(* Logix 5000 project; controller PLC_MCC1201_220AP1 vendor 1 type 14 code 164 rev 35.11; software revision 35.00; part 16 of 25 *)
(* tags used below, declared in another part *)
   AFI : ALIAS FOR B3[7].15;
   B151 : DINT[20];
   B152 : DINT[50];
   B153 : DINT[20];
   B154 : DINT[20];
   B155 : DINT[20];
   B3 : DINT[102];
   BT41_006 : MESSAGE;   // Block Transfer Read Control for Analog Input Card in Washer Panel
   BT41_007 : MESSAGE;   // Block Transfer Write Control for Analog Input Card in Washer Panel
   C1_ACK : ALIAS FOR N54[260].14;
   C1_ACTIVE_LAMP : ALIAS FOR N54[260].0;
   C1_BEACON : ALIAS FOR O[27].6;
   C1_BEACON2 : ALIAS FOR O[47].10;
   C1_HORN : ALIAS FOR O[27].5;
   C1_NTH_IN_LMP : ALIAS FOR N54[260].10;
   C1_NTH_IN_PE : ALIAS FOR N54[260].6;
   C1_NTH_IN_SS : ALIAS FOR N54[260].2;
   C1_NTH_OUT_LMP : ALIAS FOR N54[260].9;
   C1_NTH_OUT_PE : ALIAS FOR N54[260].5;
   C1_NTH_OUT_SS : ALIAS FOR N54[260].1;
   C1_STH_IN_LMP : ALIAS FOR N54[260].12;
   C1_STH_IN_PE : ALIAS FOR N54[260].8;
   C1_STH_IN_SS : ALIAS FOR N54[260].4;
   C1_STH_OUT_LMP : ALIAS FOR N54[260].11;
   C1_STH_OUT_PE : ALIAS FOR N54[260].7;
   C1_STH_OUT_SS : ALIAS FOR N54[260].3;
   C2_ACTIVE_LAMP : ALIAS FOR N54[261].0;
   C2_NTH_IN_LMP : ALIAS FOR N54[261].10;
   C2_NTH_IN_PE : ALIAS FOR N54[261].6;
   C2_NTH_IN_SS : ALIAS FOR N54[261].2;
   C2_NTH_OUT_LMP : ALIAS FOR N54[261].9;
   C2_NTH_OUT_PE : ALIAS FOR N54[261].5;
   C2_NTH_OUT_SS : ALIAS FOR N54[261].1;
   C2_STH_IN_LMP : ALIAS FOR N54[261].12;
   C2_STH_IN_PE : ALIAS FOR N54[261].8;
   C2_STH_IN_SS : ALIAS FOR N54[261].4;
   C2_STH_OUT_LMP : ALIAS FOR N54[261].11;
   C2_STH_OUT_PE : ALIAS FOR N54[261].7;
   C2_STH_OUT_SS : ALIAS FOR N54[261].3;
   C3_ACTIVE_LAMP : ALIAS FOR N54[262].0;
   C3_NTH_IN_LMP : ALIAS FOR N54[262].10;
   C3_NTH_IN_PE : ALIAS FOR N54[262].6;
   C3_NTH_IN_SS : ALIAS FOR N54[262].2;
   C3_NTH_OUT_LMP : ALIAS FOR N54[262].9;
   C3_NTH_OUT_PE : ALIAS FOR N54[262].5;
   C3_NTH_OUT_SS : ALIAS FOR N54[262].1;
   C3_STH_IN_LMP : ALIAS FOR N54[262].12;
   C3_STH_IN_PE : ALIAS FOR N54[262].8;
   C3_STH_IN_SS : ALIAS FOR N54[262].4;
   C3_STH_OUT_LMP : ALIAS FOR N54[262].11;
   C3_STH_OUT_PE : ALIAS FOR N54[262].7;
   C3_STH_OUT_SS : ALIAS FOR N54[262].3;
   C5 : COUNTER[100];
   C5_ACTIVE_LAMP : ALIAS FOR N54[264].0;
   C5_NTH_IN_LMP : ALIAS FOR N54[264].10;
   C5_NTH_IN_PE : ALIAS FOR N54[264].6;
   C5_NTH_IN_SS : ALIAS FOR N54[264].2;
   C5_NTH_OUT_LMP : ALIAS FOR N54[264].9;
   C5_NTH_OUT_PE : ALIAS FOR N54[264].5;
   C5_NTH_OUT_SS : ALIAS FOR N54[264].1;
   C5_STH_IN_LMP : ALIAS FOR N54[264].12;
   C5_STH_IN_PE : ALIAS FOR N54[264].8;
   C5_STH_IN_SS : ALIAS FOR N54[264].4;
   C5_STH_OUT_LMP : ALIAS FOR N54[264].11;
   C5_STH_OUT_PE : ALIAS FOR N54[264].7;
   C5_STH_OUT_SS : ALIAS FOR N54[264].3;
   CB_AT_SS_CUTTERS : ALIAS FOR B3[4].0;
   CR1_AUTO : ALIAS FOR I[64].13;
   CR1_DOWN_PROX : ALIAS FOR I[64].11;
   CR1_UP_PROX : ALIAS FOR I[64].12;
   F74 : REAL[2];
   F8 : REAL[20];
   I : INT[128];
   LEHR_2IN_PULSE : ALIAS FOR B73[0].1;
   M1_ALM_SILENCE : ALIAS FOR I[64].8;
   N33 : DINT[1000];
   N42 : DINT[89];
   N43 : DINT[240];
   N50 : DINT[40];
   N54 : DINT[501];
   N61 : DINT[100];
   N75 : DINT[2];
   N80 : DINT[16];
   O : INT[128];
   R150 : CONTROL[6];
   RELDR_ESTOP : ALIAS FOR I[80].0;
   Status : INT;   // INT tag to retrieve Status value through GSV created during conversion
   T4 : TIMER[100];
   T51 : TIMER[13];
   TMP_xAlwaysOFF : BOOL;
   TONY : ALIAS FOR B3[10].15;
   Z_ONS_BIT : BOOL[32];   // Temporary Boolean tag created during conversion
(* MainProgram, continued *)

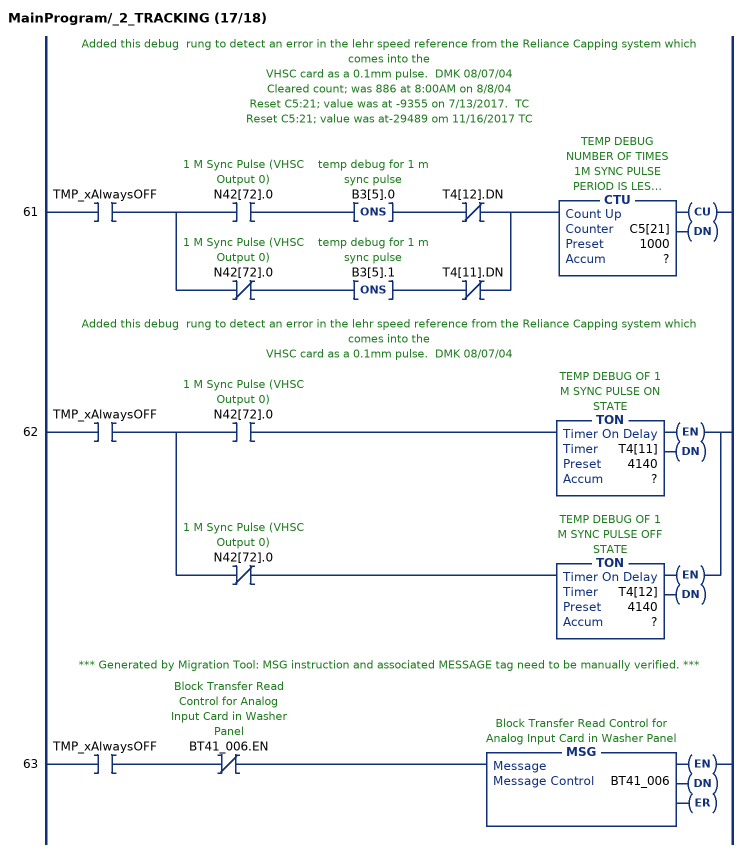
   [picture p238: MainProgram/_2_TRACKING rungs 61-63]
   // Added this debug  rung to detect an error in the lehr speed reference from the Reliance Capping system which comes into the
   // VHSC card as a 0.1mm pulse.  DMK 08/07/04
   // Cleared count; was 886 at 8:00AM on 8/8/04
   //  Reset C5:21; value was at -9355 on 7/13/2017.  TC
   // Reset C5:21; value was at-29489 om 11/16/2017 TC
   61: XIC(TMP_xAlwaysOFF)[XIC(N42[72].0) ONS(B3[5].0) XIO(T4[12].DN) ,XIO(N42[72].0) ONS(B3[5].1) XIO(T4[11].DN) ]CTU(C5[21],?,?);
   // Added this debug  rung to detect an error in the lehr speed reference from the Reliance Capping system which comes into the
   // VHSC card as a 0.1mm pulse.  DMK 08/07/04
   62: XIC(TMP_xAlwaysOFF)[XIC(N42[72].0) TON(T4[11],?,?) ,XIO(N42[72].0) TON(T4[12],?,?) ];
   // *** Generated by Migration Tool: MSG instruction and associated MESSAGE tag need to be manually verified. ***
   63: XIC(TMP_xAlwaysOFF)XIO(BT41_006.EN)MSG(BT41_006);
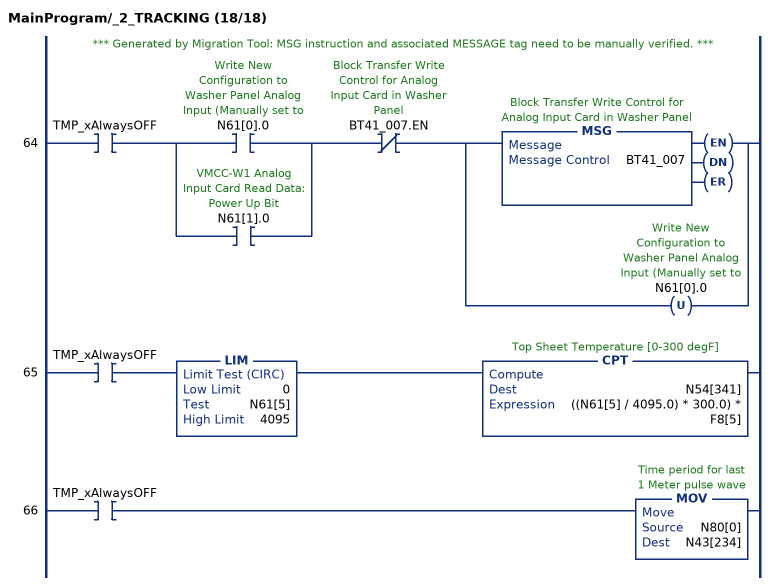
   // *** Generated by Migration Tool: MSG instruction and associated MESSAGE tag need to be manually verified. ***
   64: XIC(TMP_xAlwaysOFF)[XIC(N61[0].0) ,XIC(N61[1].0) ]XIO(BT41_007.EN)[MSG(BT41_007) ,OTU(N61[0].0) ];
   65: XIC(TMP_xAlwaysOFF)LIM(0,N61[5],4095)CPT(N54[341],((N61[5] / 4095.0) * 300.0) * F8[5]);
   66: XIC(TMP_xAlwaysOFF)MOV(N80[0],N43[234]);
END_ROUTINE

ROUTINE _31_MSEC   (* ladder *)
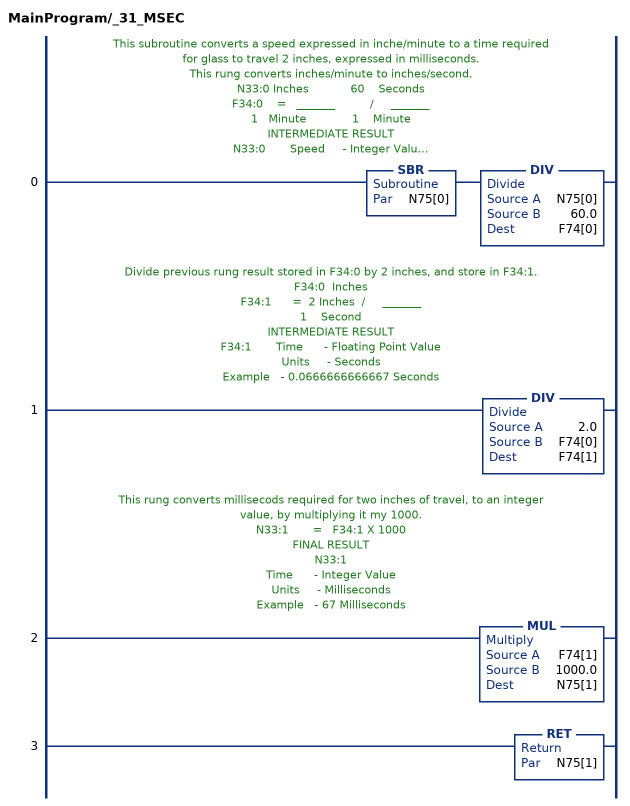
   // This subroutine converts a speed expressed in inche/minute to a time required
   // for glass to travel 2 inches, expressed in milliseconds.
   // This rung converts inches/minute to inches/second.
   //                    N33:0 Inches            60    Seconds
   //      F34:0    =   _______          /     _______
   //                      1   Minute             1    Minute
   // INTERMEDIATE RESULT
   // N33:0       Speed     - Integer Value
   //             Units     - Inches / Minute
   //             Example   - 1800 Inches / Minute
   // F34:0       Speed     - Floating Point Value
   //             Units     - Inches / Second
   //             Example   - 30 Inches / Second
   // HISTORY
   // DATE        DESCRIPTION                                               PROGRAMMER
   // ----        -----------                                               ----------
   // 11/93       Subroutine created for Lathrop MAIN_3 5/40 processor.     WAS
   // 3/11/95     Subroutine imported, addresses changed.                   WAS
   // 1/29/96     Imported subroutine into Laurinburg processor MB for
   //             75F1 marking bridge/front end PLC control. Will use for
   //             tracking crossbreaks.                                     WAS
   0: SBR(N75[0])DIV(N75[0],60.0,F74[0]);
   // Divide previous rung result stored in F34:0 by 2 inches, and store in F34:1.
   //                                     F34:0  Inches
   //      F34:1      =  2 Inches  /     _______
   //                                       1    Second
   // INTERMEDIATE RESULT
   // F34:1       Time      - Floating Point Value
   //             Units     - Seconds
   //             Example   - 0.0666666666667 Seconds
   1: DIV(2.0,F74[0],F74[1]);
   // This rung converts millisecods required for two inches of travel, to an integer
   //  value, by multiplying it my 1000.
   // N33:1       =   F34:1 X 1000
   // FINAL RESULT
   // N33:1
   //             Time      - Integer Value
   //             Units     - Milliseconds
   //             Example   - 67 Milliseconds
   2: MUL(F74[1],1000.0,N75[1]);
   3: RET(N75[1]);
END_ROUTINE

ROUTINE _41_C1_OPS   (* ladder *)
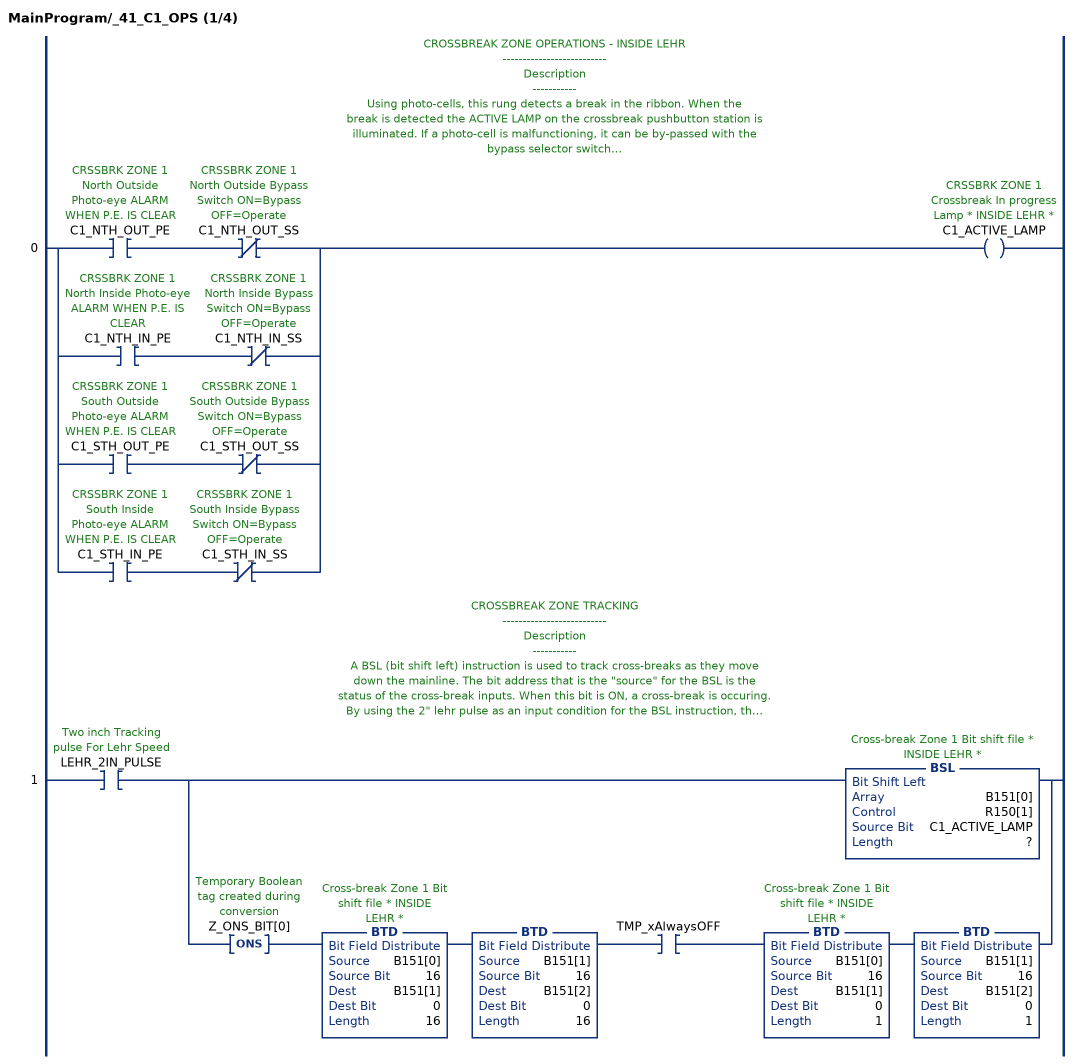
   // CROSSBREAK ZONE OPERATIONS - INSIDE LEHR
   // --------------------------
   // Description
   // -----------
   // Using photo-cells, this rung detects a break in the ribbon. When the
   // break is detected the ACTIVE LAMP on the crossbreak pushbutton station is
   // illuminated. If a photo-cell is malfunctioning, it can be by-passed with the
   // bypass selector switch.
   // History
   // =======
   // DATE        DESCRIPTION                                               PROGRAMMER
   // ----        -----------                                               ----------
   // 1/22/96     Created cross-break rungs, imported symbols and coil      WAS
   //             comments from MS-Excel CSV file, and placed comments
   //             for each rung.
   0: [XIC(C1_NTH_OUT_PE) XIO(C1_NTH_OUT_SS) ,XIC(C1_NTH_IN_PE) XIO(C1_NTH_IN_SS) ,XIC(C1_STH_OUT_PE) XIO(C1_STH_OUT_SS) ,XIC(C1_STH_IN_PE) XIO(C1_STH_IN_SS) ]OTE(C1_ACTIVE_LAMP);
   // CROSSBREAK ZONE TRACKING
   // --------------------------
   // Description
   // -----------
   // A BSL (bit shift left) instruction is used to track cross-breaks as they move
   // down the mainline. The bit address that is the "source" for the BSL is the
   // status of the cross-break inputs. When this bit is ON, a cross-break is occuring.
   // By using the 2" lehr pulse as an input condition for the BSL instruction, the
   // cross-break information is shifted to track the movement of the ribbon.
   // History
   // =======
   // DATE        DESCRIPTION                                               PROGRAMMER
   // ----        -----------                                               ----------
   // 1/30/96     Entered BSL instructions for all cross-break zones        WAS
   1: XIC(LEHR_2IN_PULSE)[BSL(B151[0],R150[1],C1_ACTIVE_LAMP,?) ,ONS(Z_ONS_BIT[0]) BTD(B151[0],16,B151[1],0,16) BTD(B151[1],16,B151[2],0,16) XIC(TMP_xAlwaysOFF) BTD(B151[0],16,B151[1],0,1) BTD(B151[1],16,B151[2],0,1) ];
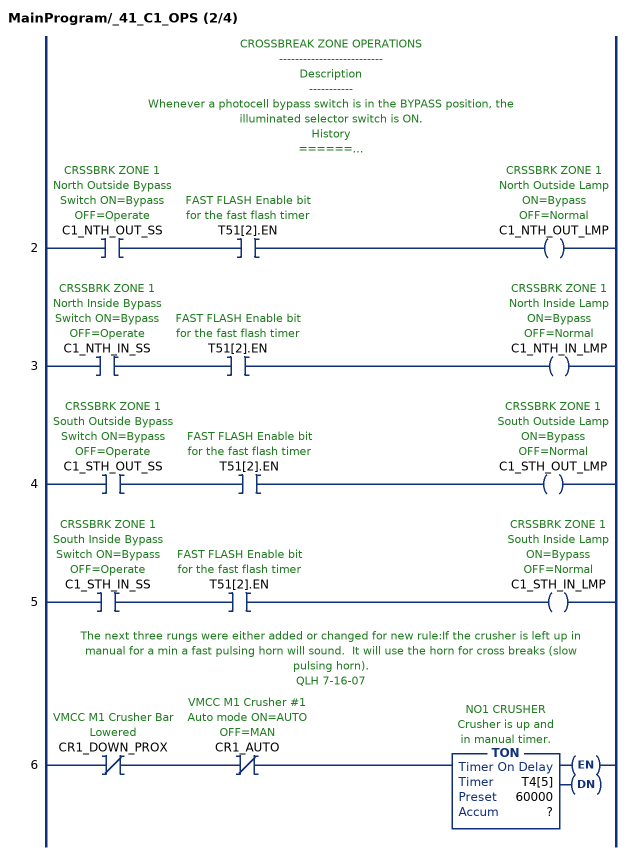
   // CROSSBREAK ZONE OPERATIONS
   // --------------------------
   // Description
   // -----------
   // Whenever a photocell bypass switch is in the BYPASS position, the
   // illuminated selector switch is ON.
   // History
   // =======
   // DATE        DESCRIPTION                                               PROGRAMMER
   // ----        -----------                                               ----------
   // 1/22/96     Created cross-break rungs, imported symbols and coil      WAS
   //             comments from MS-Excel CSV file, and placed comments
   //             for each rung.
   2: XIC(C1_NTH_OUT_SS)XIC(T51[2].EN)OTE(C1_NTH_OUT_LMP);
   3: XIC(C1_NTH_IN_SS)XIC(T51[2].EN)OTE(C1_NTH_IN_LMP);
   4: XIC(C1_STH_OUT_SS)XIC(T51[2].EN)OTE(C1_STH_OUT_LMP);
   5: XIC(C1_STH_IN_SS)XIC(T51[2].EN)OTE(C1_STH_IN_LMP);
   // The next three rungs were either added or changed for new rule:If the crusher is left up in manual for a min a fast pulsing horn will sound.  It will use the horn for cross breaks (slow pulsing horn).
   // QLH 7-16-07
   6: XIO(CR1_DOWN_PROX)XIO(CR1_AUTO)TON(T4[5],?,?);
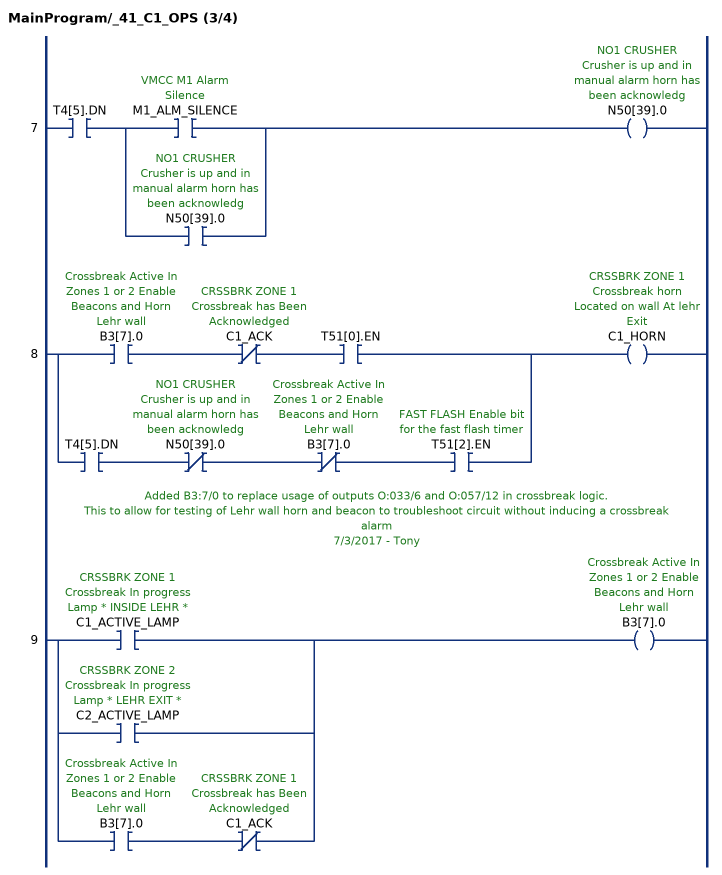
   7: XIC(T4[5].DN)[XIC(M1_ALM_SILENCE) ,XIC(N50[39].0) ]OTE(N50[39].0);
   8: [XIC(B3[7].0) XIO(C1_ACK) XIC(T51[0].EN) ,XIC(T4[5].DN) XIO(N50[39].0) XIO(B3[7].0) XIC(T51[2].EN) ]OTE(C1_HORN);
   // Added B3:7/0 to replace usage of outputs O:033/6 and O:057/12 in crossbreak logic.
   //                                                                         This to allow for testing of Lehr wall horn and beacon to troubleshoot circuit without inducing a crossbreak alarm
   //                                                                                                                                          7/3/2017 - Tony
   9: [[XIC(C1_ACTIVE_LAMP) ,XIC(C2_ACTIVE_LAMP) ] ,XIC(B3[7].0) XIO(C1_ACK) ]OTE(B3[7].0);
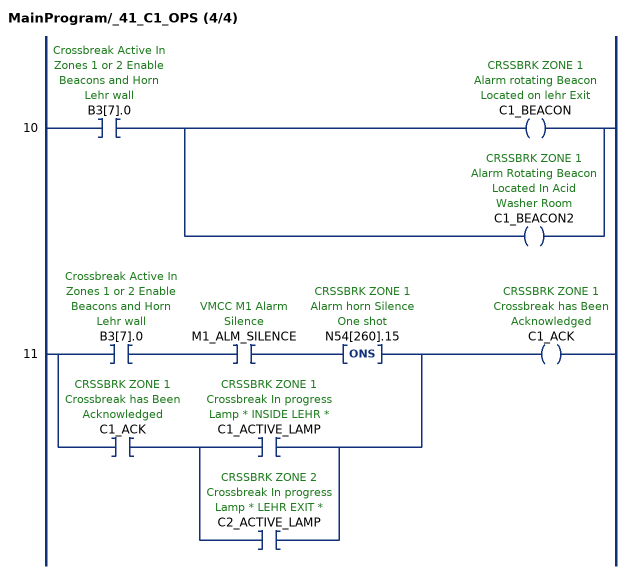
   10: XIC(B3[7].0)[OTE(C1_BEACON) ,OTE(C1_BEACON2) ];
   11: [XIC(B3[7].0) XIC(M1_ALM_SILENCE) ONS(N54[260].15) ,XIC(C1_ACK) [XIC(C1_ACTIVE_LAMP) ,XIC(C2_ACTIVE_LAMP) ] ]OTE(C1_ACK);
END_ROUTINE

ROUTINE _42_C2_OPS   (* ladder *)
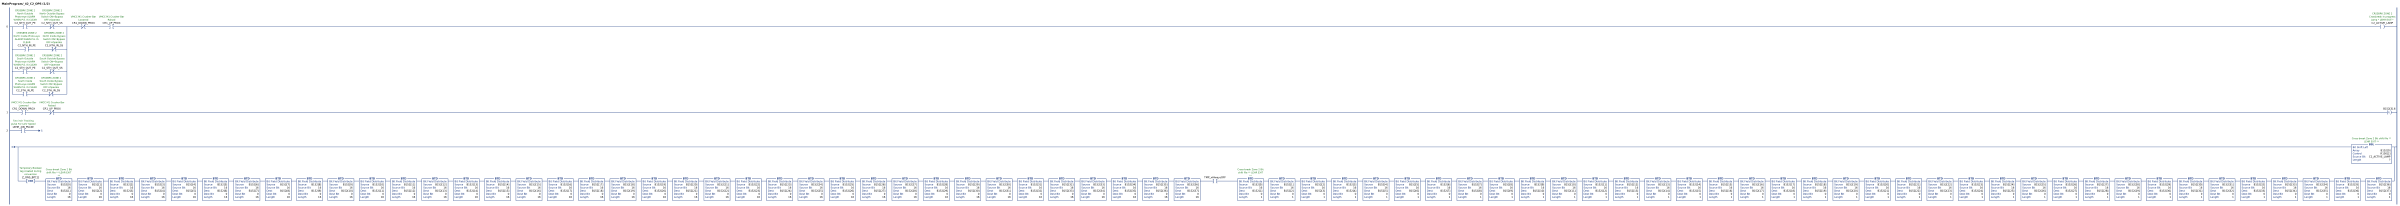
   0: [XIC(C2_NTH_OUT_PE) XIO(C2_NTH_OUT_SS) ,XIC(C2_NTH_IN_PE) XIO(C2_NTH_IN_SS) ,XIC(C2_STH_OUT_PE) XIO(C2_STH_OUT_SS) ,XIC(C2_STH_IN_PE) XIO(C2_STH_IN_SS) ]XIO(CR1_DOWN_PROX)XIC(CR1_UP_PROX)OTE(C2_ACTIVE_LAMP);
   1: XIC(CR1_DOWN_PROX)XIO(CR1_UP_PROX)OTL(B152[3].6);
   2: XIC(LEHR_2IN_PULSE)[BSL(B152[0],R150[2],C2_ACTIVE_LAMP,?) ,ONS(Z_ONS_BIT[1]) BTD(B152[0],16,B152[1],0,16) BTD(B152[1],16,B152[2],0,16) BTD(B152[2],16,B152[3],0,16) BTD(B152[3],16,B152[4],0,16) BTD(B152[4],16,B152[5],0,16) BTD(B152[5],16,B152[6],0,16) BTD(B152[6],16,B152[7],0,16) BTD(B152[7],16,B152[8],0,16) BTD(B152[8],16,B152[9],0,16) BTD(B152[9],16,B152[10],0,16) BTD(B152[10],16,B152[11],0,16) BTD(B152[11],16,B152[12],0,16) BTD(B152[12],16,B152[13],0,16) BTD(B152[13],16,B152[14],0,16) BTD(B152[14],16,B152[15],0,16) BTD(B152[15],16,B152[16],0,16) BTD(B152[16],16,B152[17],0,16) BTD(B152[17],16,B152[18],0,16) BTD(B152[18],16,B152[19],0,16) BTD(B152[19],16,B152[20],0,16) BTD(B152[20],16,B152[21],0,16) BTD(B152[21],16,B152[22],0,16) BTD(B152[22],16,B152[23],0,16) BTD(B152[23],16,B152[24],0,16) BTD(B152[24],16,B152[25],0,16) BTD(B152[25],16,B152[26],0,16) BTD(B152[26],16,B152[27],0,16) BTD(B152[27],16,B152[28],0,16) BTD(B152[28],16,B152[29],0,16) BTD(B152[29],16,B152[30],0,16) BTD(B152[30],16,B152[31],0,16) BTD(B152[31],16,B152[32],0,16) BTD(B152[32],16,B152[33],0,16) BTD(B152[33],16,B152[34],0,16) BTD(B152[34],16,B152[35],0,16) BTD(B152[35],16,B152[36],0,16) BTD(B152[36],16,B152[37],0,16) XIC(TMP_xAlwaysOFF) BTD(B152[0],16,B152[1],0,1) BTD(B152[1],16,B152[2],0,1) BTD(B152[2],16,B152[3],0,1) BTD(B152[3],16,B152[4],0,1) BTD(B152[4],16,B152[5],0,1) BTD(B152[5],16,B152[6],0,1) BTD(B152[6],16,B152[7],0,1) BTD(B152[7],16,B152[8],0,1) BTD(B152[8],16,B152[9],0,1) BTD(B152[9],16,B152[10],0,1) BTD(B152[10],16,B152[11],0,1) BTD(B152[11],16,B152[12],0,1) BTD(B152[12],16,B152[13],0,1) BTD(B152[13],16,B152[14],0,1) BTD(B152[14],16,B152[15],0,1) BTD(B152[15],16,B152[16],0,1) BTD(B152[16],16,B152[17],0,1) BTD(B152[17],16,B152[18],0,1) BTD(B152[18],16,B152[19],0,1) BTD(B152[19],16,B152[20],0,1) BTD(B152[20],16,B152[21],0,1) BTD(B152[21],16,B152[22],0,1) BTD(B152[22],16,B152[23],0,1) BTD(B152[23],16,B152[24],0,1) BTD(B152[24],16,B152[25],0,1) BTD(B152[25],16,B152[26],0,1) BTD(B152[26],16,B152[27],0,1) BTD(B152[27],16,B152[28],0,1) BTD(B152[28],16,B152[29],0,1) BTD(B152[29],16,B152[30],0,1) BTD(B152[30],16,B152[31],0,1) BTD(B152[31],16,B152[32],0,1) BTD(B152[32],16,B152[33],0,1) BTD(B152[33],16,B152[34],0,1) BTD(B152[34],16,B152[35],0,1) BTD(B152[35],16,B152[36],0,1) BTD(B152[36],16,B152[37],0,1) ];
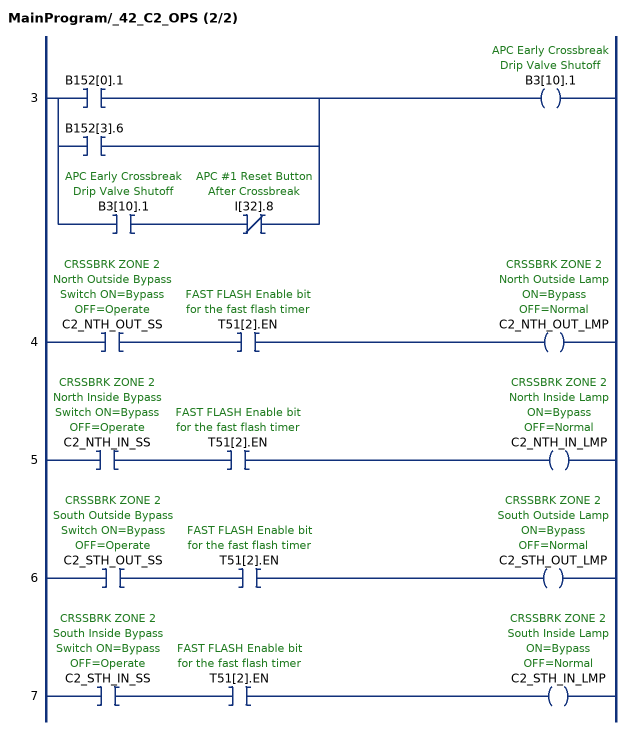
   3: [XIC(B152[0].1) ,XIC(B152[3].6) ,XIC(B3[10].1) XIO(I[32].8) ]OTE(B3[10].1);
   4: XIC(C2_NTH_OUT_SS)XIC(T51[2].EN)OTE(C2_NTH_OUT_LMP);
   5: XIC(C2_NTH_IN_SS)XIC(T51[2].EN)OTE(C2_NTH_IN_LMP);
   6: XIC(C2_STH_OUT_SS)XIC(T51[2].EN)OTE(C2_STH_OUT_LMP);
   7: XIC(C2_STH_IN_SS)XIC(T51[2].EN)OTE(C2_STH_IN_LMP);
END_ROUTINE

ROUTINE _43_C3_OPS   (* ladder *)
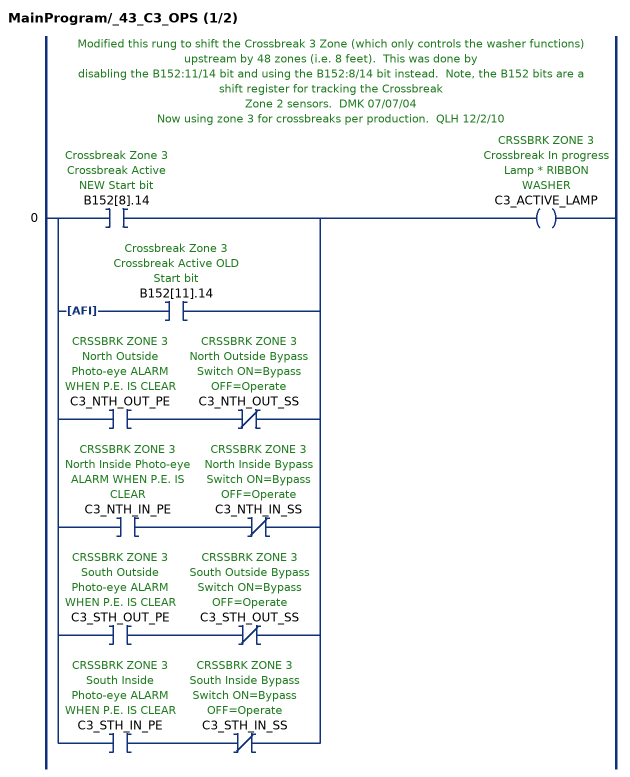
   // Modified this rung to shift the Crossbreak 3 Zone (which only controls the washer functions) upstream by 48 zones (i.e. 8 feet).  This was done by
   // disabling the B152:11/14 bit and using the B152:8/14 bit instead.  Note, the B152 bits are a shift register for tracking the Crossbreak
   // Zone 2 sensors.  DMK 07/07/04
   // Now using zone 3 for crossbreaks per production.  QLH 12/2/10
   0: [XIC(B152[8].14) ,AFI() XIC(B152[11].14) ,XIC(C3_NTH_OUT_PE) XIO(C3_NTH_OUT_SS) ,XIC(C3_NTH_IN_PE) XIO(C3_NTH_IN_SS) ,XIC(C3_STH_OUT_PE) XIO(C3_STH_OUT_SS) ,XIC(C3_STH_IN_PE) XIO(C3_STH_IN_SS) ]OTE(C3_ACTIVE_LAMP);
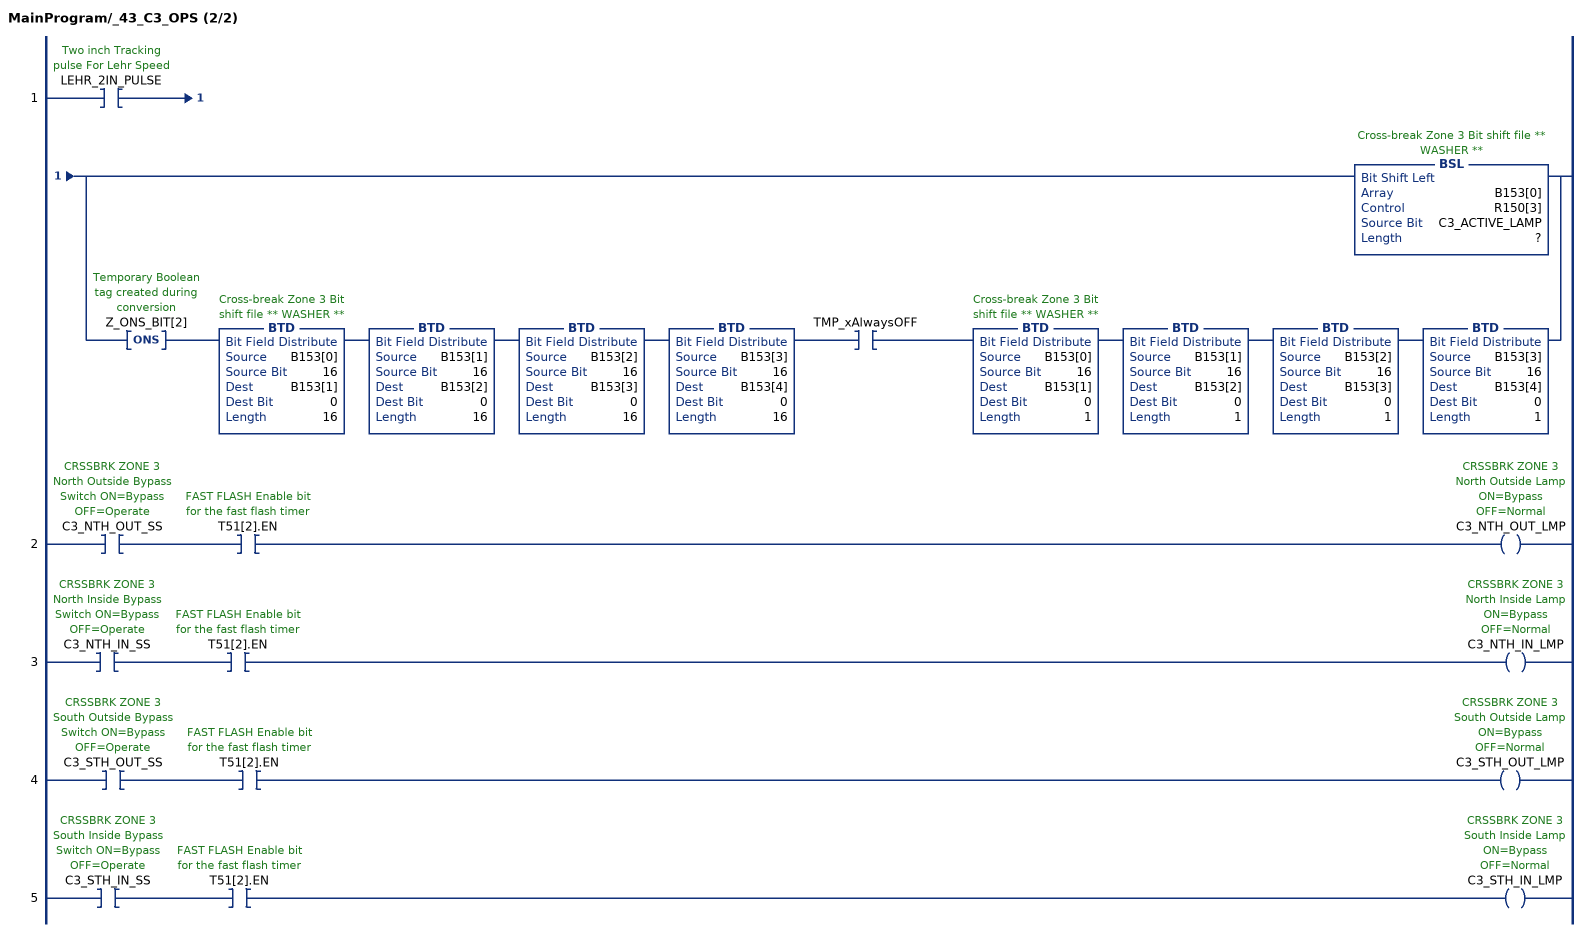
   1: XIC(LEHR_2IN_PULSE)[BSL(B153[0],R150[3],C3_ACTIVE_LAMP,?) ,ONS(Z_ONS_BIT[2]) BTD(B153[0],16,B153[1],0,16) BTD(B153[1],16,B153[2],0,16) BTD(B153[2],16,B153[3],0,16) BTD(B153[3],16,B153[4],0,16) XIC(TMP_xAlwaysOFF) BTD(B153[0],16,B153[1],0,1) BTD(B153[1],16,B153[2],0,1) BTD(B153[2],16,B153[3],0,1) BTD(B153[3],16,B153[4],0,1) ];
   2: XIC(C3_NTH_OUT_SS)XIC(T51[2].EN)OTE(C3_NTH_OUT_LMP);
   3: XIC(C3_NTH_IN_SS)XIC(T51[2].EN)OTE(C3_NTH_IN_LMP);
   4: XIC(C3_STH_OUT_SS)XIC(T51[2].EN)OTE(C3_STH_OUT_LMP);
   5: XIC(C3_STH_IN_SS)XIC(T51[2].EN)OTE(C3_STH_IN_LMP);
END_ROUTINE

ROUTINE _44_LADDER   (* ladder *)
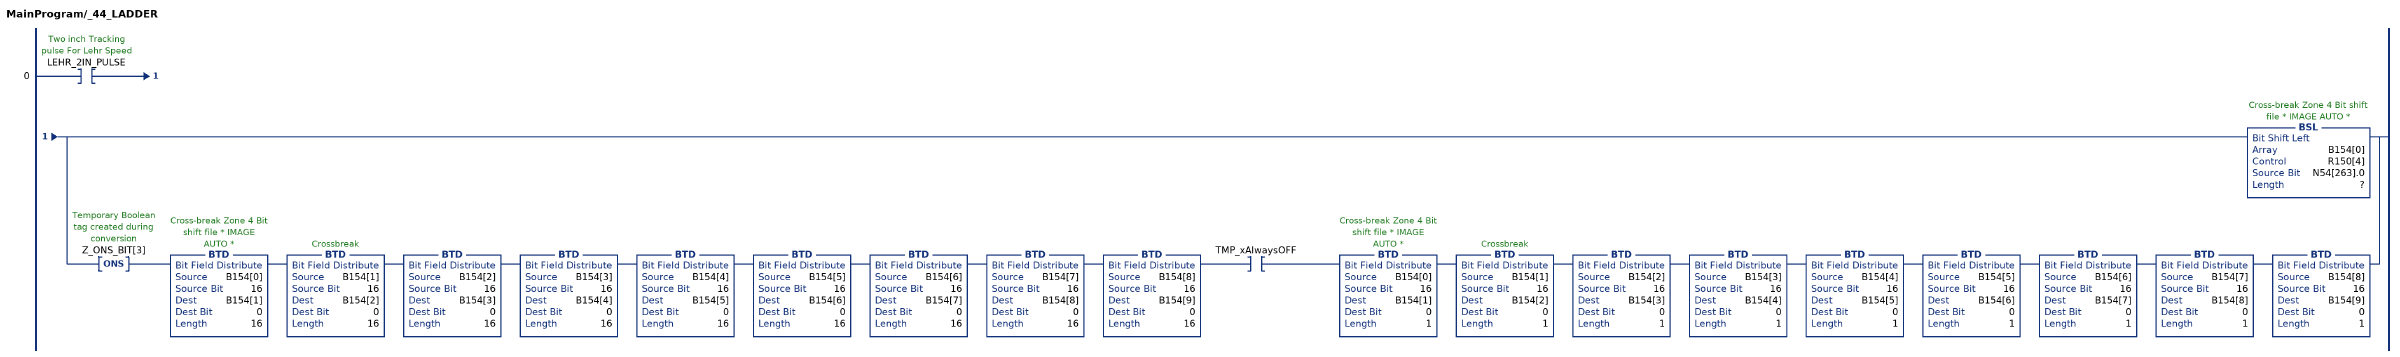
   0: XIC(LEHR_2IN_PULSE)[BSL(B154[0],R150[4],N54[263].0,?) ,ONS(Z_ONS_BIT[3]) BTD(B154[0],16,B154[1],0,16) BTD(B154[1],16,B154[2],0,16) BTD(B154[2],16,B154[3],0,16) BTD(B154[3],16,B154[4],0,16) BTD(B154[4],16,B154[5],0,16) BTD(B154[5],16,B154[6],0,16) BTD(B154[6],16,B154[7],0,16) BTD(B154[7],16,B154[8],0,16) BTD(B154[8],16,B154[9],0,16) XIC(TMP_xAlwaysOFF) BTD(B154[0],16,B154[1],0,1) BTD(B154[1],16,B154[2],0,1) BTD(B154[2],16,B154[3],0,1) BTD(B154[3],16,B154[4],0,1) BTD(B154[4],16,B154[5],0,1) BTD(B154[5],16,B154[6],0,1) BTD(B154[6],16,B154[7],0,1) BTD(B154[7],16,B154[8],0,1) BTD(B154[8],16,B154[9],0,1) ];
END_ROUTINE

ROUTINE _45_C5_OPS   (* ladder *)
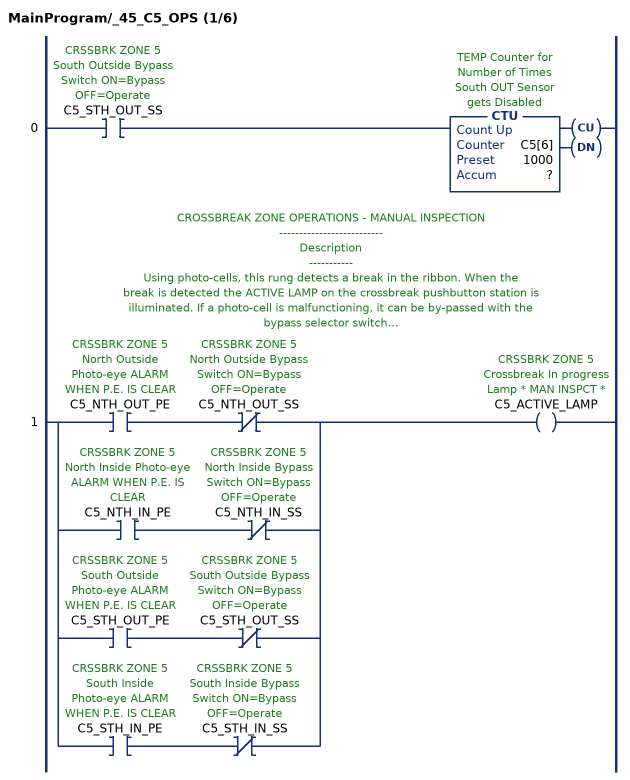
   0: XIC(C5_STH_OUT_SS)CTU(C5[6],?,?);
   // CROSSBREAK ZONE OPERATIONS - MANUAL INSPECTION
   // --------------------------
   // Description
   // -----------
   // Using photo-cells, this rung detects a break in the ribbon. When the
   // break is detected the ACTIVE LAMP on the crossbreak pushbutton station is
   // illuminated. If a photo-cell is malfunctioning, it can be by-passed with the
   // bypass selector switch.
   // History
   // =======
   // DATE        DESCRIPTION
   // PROGRAMMER
   // ----        -----------
   // ----------
   // 1/22/96     Created cross-break rungs, imported symbols and coil      WAS
   //             comments from MS-Excel CSV file, and placed comments
   //             for each rung.
   1: [XIC(C5_NTH_OUT_PE) XIO(C5_NTH_OUT_SS) ,XIC(C5_NTH_IN_PE) XIO(C5_NTH_IN_SS) ,XIC(C5_STH_OUT_PE) XIO(C5_STH_OUT_SS) ,XIC(C5_STH_IN_PE) XIO(C5_STH_IN_SS) ]OTE(C5_ACTIVE_LAMP);
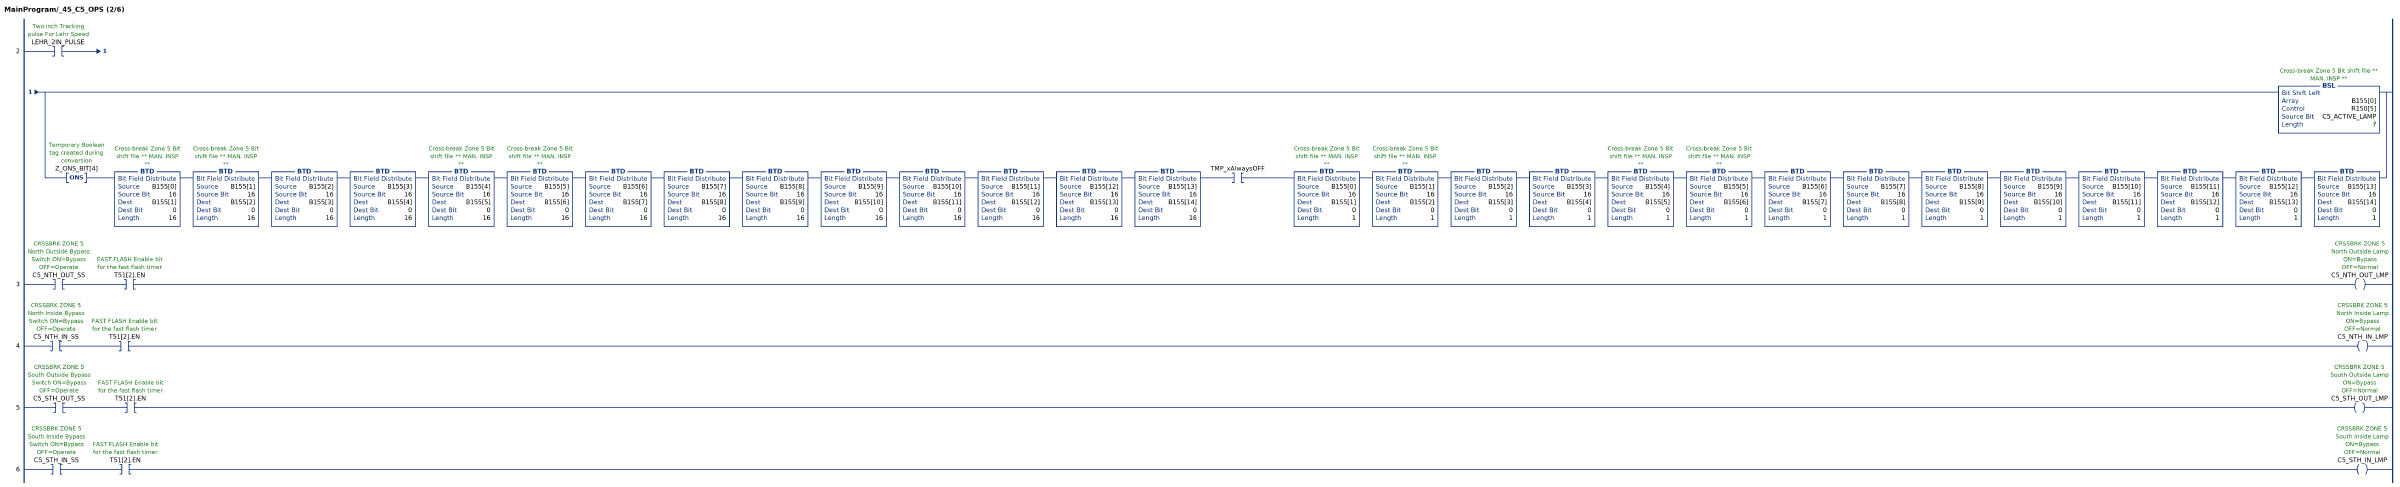
   2: XIC(LEHR_2IN_PULSE)[BSL(B155[0],R150[5],C5_ACTIVE_LAMP,?) ,ONS(Z_ONS_BIT[4]) BTD(B155[0],16,B155[1],0,16) BTD(B155[1],16,B155[2],0,16) BTD(B155[2],16,B155[3],0,16) BTD(B155[3],16,B155[4],0,16) BTD(B155[4],16,B155[5],0,16) BTD(B155[5],16,B155[6],0,16) BTD(B155[6],16,B155[7],0,16) BTD(B155[7],16,B155[8],0,16) BTD(B155[8],16,B155[9],0,16) BTD(B155[9],16,B155[10],0,16) BTD(B155[10],16,B155[11],0,16) BTD(B155[11],16,B155[12],0,16) BTD(B155[12],16,B155[13],0,16) BTD(B155[13],16,B155[14],0,16) XIC(TMP_xAlwaysOFF) BTD(B155[0],16,B155[1],0,1) BTD(B155[1],16,B155[2],0,1) BTD(B155[2],16,B155[3],0,1) BTD(B155[3],16,B155[4],0,1) BTD(B155[4],16,B155[5],0,1) BTD(B155[5],16,B155[6],0,1) BTD(B155[6],16,B155[7],0,1) BTD(B155[7],16,B155[8],0,1) BTD(B155[8],16,B155[9],0,1) BTD(B155[9],16,B155[10],0,1) BTD(B155[10],16,B155[11],0,1) BTD(B155[11],16,B155[12],0,1) BTD(B155[12],16,B155[13],0,1) BTD(B155[13],16,B155[14],0,1) ];
   3: XIC(C5_NTH_OUT_SS)XIC(T51[2].EN)OTE(C5_NTH_OUT_LMP);
   4: XIC(C5_NTH_IN_SS)XIC(T51[2].EN)OTE(C5_NTH_IN_LMP);
   5: XIC(C5_STH_OUT_SS)XIC(T51[2].EN)OTE(C5_STH_OUT_LMP);
   6: XIC(C5_STH_IN_SS)XIC(T51[2].EN)OTE(C5_STH_IN_LMP);
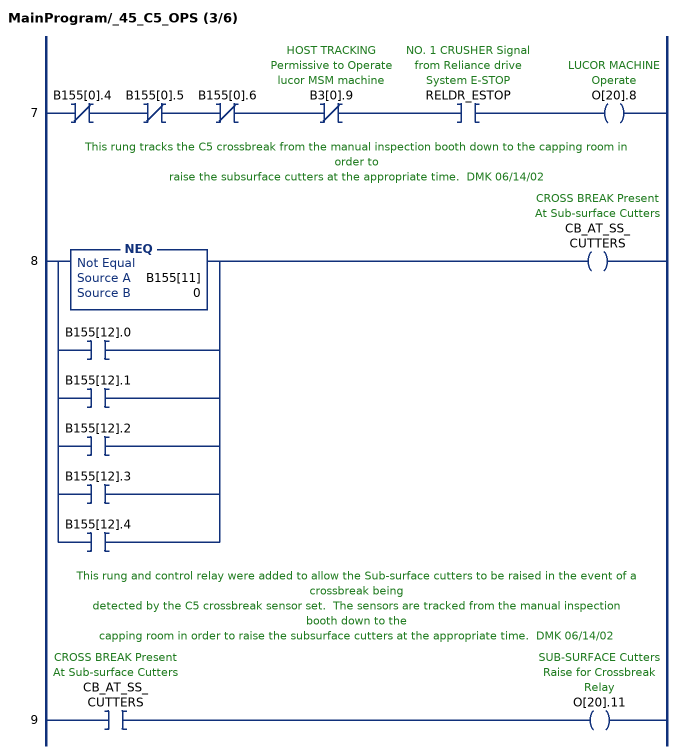
   7: XIO(B155[0].4)XIO(B155[0].5)XIO(B155[0].6)XIO(B3[0].9)XIC(RELDR_ESTOP)OTE(O[20].8);
   // This rung tracks the C5 crossbreak from the manual inspection booth down to the capping room in order to
   // raise the subsurface cutters at the appropriate time.  DMK 06/14/02
   8: [NEQ(B155[11],0) ,XIC(B155[12].0) ,XIC(B155[12].1) ,XIC(B155[12].2) ,XIC(B155[12].3) ,XIC(B155[12].4) ]OTE(CB_AT_SS_CUTTERS);
   // This rung and control relay were added to allow the Sub-surface cutters to be raised in the event of a crossbreak being
   // detected by the C5 crossbreak sensor set.  The sensors are tracked from the manual inspection booth down to the
   // capping room in order to raise the subsurface cutters at the appropriate time.  DMK 06/14/02
   9: XIC(CB_AT_SS_CUTTERS)OTE(O[20].11);
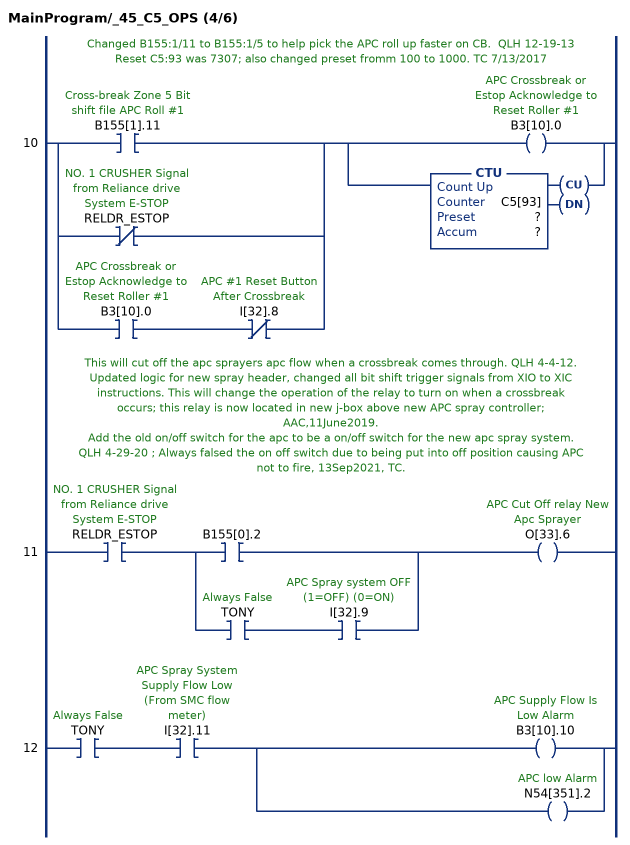
   // Changed B155:1/11 to B155:1/5 to help pick the APC roll up faster on CB.  QLH 12-19-13
   // Reset C5:93 was 7307; also changed preset fromm 100 to 1000. TC 7/13/2017
   10: [[XIC(B155[1].11) ,XIO(RELDR_ESTOP) ] ,XIC(B3[10].0) XIO(I[32].8) ][OTE(B3[10].0) ,CTU(C5[93],?,?) ];
   // This will cut off the apc sprayers apc flow when a crossbreak comes through. QLH 4-4-12.
   //                                              Updated logic for new spray header, changed all bit shift trigger signals from XIO to XIC instructions. This will change the operation of the relay to turn on when a crossbreak occurs; this relay is now located in new j-box above new APC spray controller; AAC,11June2019.
   //                                              Add the old on/off switch for the apc to be a on/off switch for the new apc spray system. QLH 4-29-20 ; Always falsed the on off switch due to being put into off position causing APC not to fire, 13Sep2021, TC.
   11: XIC(RELDR_ESTOP)[XIC(B155[0].2) ,XIC(TONY) XIC(I[32].9) ]OTE(O[33].6);
   12: XIC(TONY)XIC(I[32].11)[OTE(B3[10].10) ,OTE(N54[351].2) ];
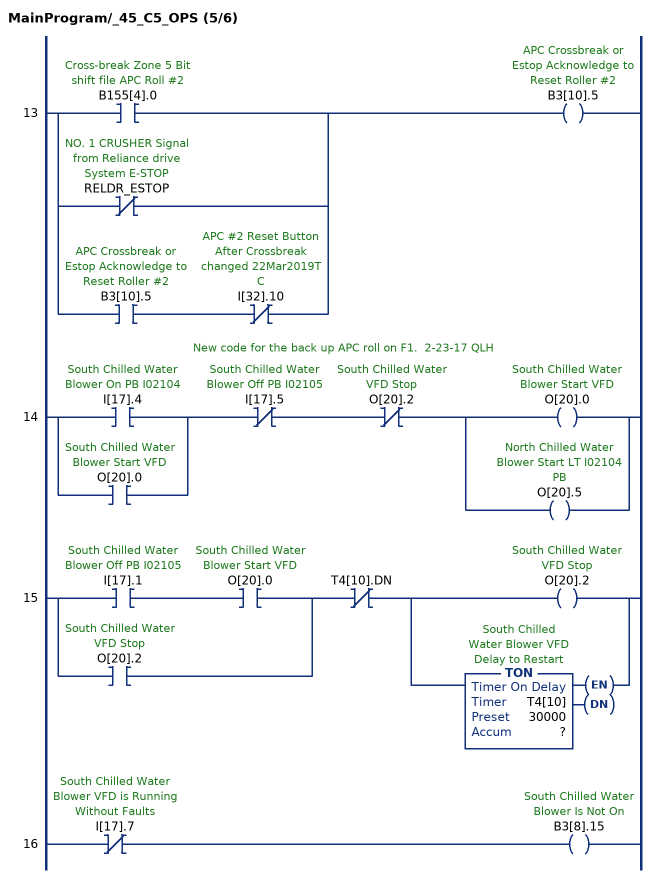
   13: [[XIC(B155[4].0) ,XIO(RELDR_ESTOP) ] ,XIC(B3[10].5) XIO(I[32].10) ]OTE(B3[10].5);
   // New code for the back up APC roll on F1.  2-23-17 QLH
   14: [XIC(I[17].4) ,XIC(O[20].0) ]XIO(I[17].5)XIO(O[20].2)[OTE(O[20].0) ,OTE(O[20].5) ];
   15: [XIC(I[17].1) XIC(O[20].0) ,XIC(O[20].2) ]XIO(T4[10].DN)[OTE(O[20].2) ,TON(T4[10],?,?) ];
   16: XIO(I[17].7)OTE(B3[8].15);
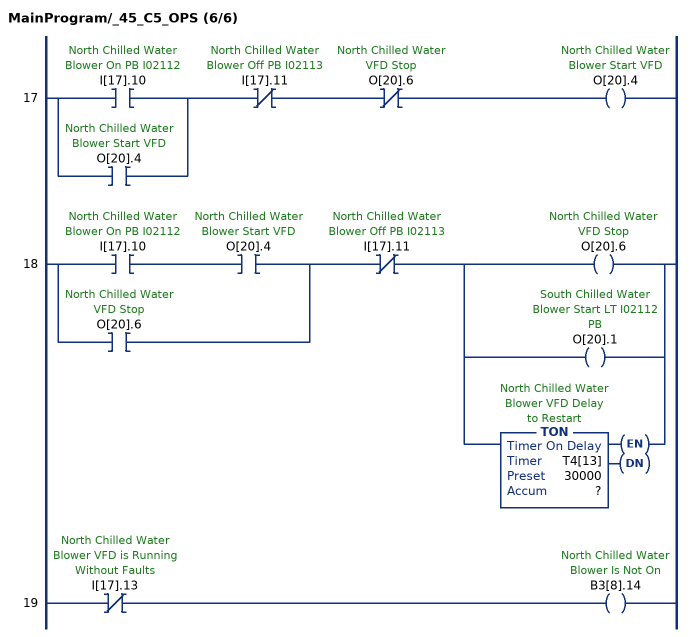
   17: [XIC(I[17].10) ,XIC(O[20].4) ]XIO(I[17].11)XIO(O[20].6)OTE(O[20].4);
   18: [XIC(I[17].10) XIC(O[20].4) ,XIC(O[20].6) ]XIO(I[17].11)[[OTE(O[20].6) ,OTE(O[20].1) ] ,TON(T4[13],?,?) ];
   19: XIO(I[17].13)OTE(B3[8].14);
END_ROUTINE
